(* Logix 5000 project; controller PLC_MCC1300_75F1 vendor 1 type 14 code 166 rev 32.11; software revision 32.04; part 3 of 83 *)
(* tags used below, declared in another part *)
   O : INT[128];
   Z301 : MAC_Zone_ML;

TYPE MAC_TrimmingWheels_PH :
STRUCT
   x0 : BOOL;   // Arming
   x1 : BOOL;
   x2 : BOOL;
   x3 : BOOL;   // Firing operator side
   x4 : BOOL;
   x5 : BOOL;
   x6 : BOOL;   // Firing opposite operator side
   x7 : BOOL;
   x8 : BOOL;
   x9 : BOOL;   // End arming
   x10 : BOOL;
   x11 : BOOL;
   x12 : BOOL;   // End firing
   x13 : BOOL;
   x14 : BOOL;
   x15 : BOOL;   // Stop conveyor request
   x16 : BOOL;
   x17 : BOOL;
   x18 : BOOL;
   x19 : BOOL;
   x20 : BOOL;   // Request position to target
   x21 : BOOL;
   x22 : BOOL;
   x23 : BOOL;   // End position
   x24 : BOOL;
   x25 : BOOL;
   x26 : BOOL;
   x27 : BOOL;
   x28 : BOOL;
   x29 : BOOL;
   x30 : BOOL;
   x31 : BOOL;
END_STRUCT
END_TYPE

TYPE MAC_Zone :
STRUCT
   ST_xConditionOKStopCycle : BOOL;   // Condition OK for stop cycle
   ST_xStartCycleRequest : BOOL;   // Start cycle request
   ST_xCycleON : BOOL;   // Cycle ON
   ST_xStopCycleRequest : BOOL;   // Stop cycle request
   ST_xStopCycleAccepted : BOOL;   // Stop cycle accepted
   ST_xStopCycleReqForAlarms : BOOL;   // Stop cycle request for emergency alarms
   ST_xStopCycleAcptForAlarms : BOOL;   // Stop cycle accepted for emergency alarms
   ST_xConveyorsNotOK : BOOL;   // Conveyors not OK
   ST_xConditionOkPhaseAdvancement : BOOL;   // Condition OK phases advancement
   ST_xConditionOkCycleON : BOOL;   // Condition OK cycle ON
   ST_xConditionOkManualMode : BOOL;   // Condition ok for manual mode
   ST_xCleaningConditionOK : BOOL;   // Cleaning condition OK
   ST_xReqCleaning : BOOL;   // Request cleaning
   ST_xCleaningAccepted : BOOL;   // Cleaning accepted
   ST_xManualModeAccepted : BOOL;   // Manual mode accepted
   ST_xManualModeRequest : BOOL;   // Manual mode request
   ST_xAutoModeAccepted : BOOL;   // Auto mode accepted
   ST_xSelectionManualMode : BOOL;   // Selection manual mode
   ST_xSelectionAutomaticMode : BOOL;   // Selection automatic mode
   ST_xEnableControlError : BOOL;   // Enable control error
   ST_xZoneError : BOOL;   // Zone error
   ST_xAlarmOff : BOOL;   // Alarm OFF
   OSR_xStartCycle : BOOL;   // OSR Start cycle
   OSR_xStopCycle : BOOL;   // OSR Stop cycle
   OSR_xForceStopCycle : BOOL;   // OSR Force stop cycle
   OSR_xAlarmAcoustic : BOOL;   // OSR Alarm acoustic
   OSR_xAlarmMuting : BOOL;   // OSR Alarm muting
   OSR_xAutomaticMode : BOOL;   // OSR Automation mode
   OS_xStartCycle : BOOL;   // OS Start cycle
   OS_xStopCycle : BOOL;   // OS Stop cycle
   OS_xForceStopCycle : BOOL;   // OS Force stop cycle
   OS_xAlarmAcoustic : BOOL;   // OS Alarm acoustic
   OS_xAlarmMuting : BOOL;   // OS Alarm muting
   OS_xAutomaticMode : BOOL;   // OS Automatic mode
   AUX_dSpeedStandby_mm_min : DINT;   // Conveyor speed in stanby [mm/min] (#COSTANT#)
   AUX_dSpeedTINUnload_mm_min : DINT;   // Conveyor speed with stacker in TIM mode [mm/min] (#COSTANT#)
   AUX_dProgressiveID : DINT;   // Progressive ID
   tmON_ResetAlarm : TIMER;   // Reset alarm
   tmON_24Vdc : TIMER;   // Presence 24Vdc timer
   tmON_400Vca : TIMER;   // Presence 400Vca timer
   tmON_EmergencyOK : TIMER;   // Emergency OK timer
   tmON_Cycle : TIMER;   // Cycle ON timer
   tmON_ForceStop : TIMER;   // Force stop cycle timer
   tmON_AllowStopCleaning : TIMER;   // Allow stop cleaning timer
   tmON_CycleAcousticAlarm : TIMER;   // Cycle acoustic alarm timer
END_STRUCT
END_TYPE

TYPE MAC_Zone_ALM :
STRUCT
   rgxEmergency : DINT[3];   // Emergency
   rgxStoppingFault : DINT[1];   // Stopping faults
   rgxFault : DINT[1];   // Faults
   rgxWarning : DINT[2];   // Warning
   rgdFaultCode : DINT[1];   // Fault codes
END_STRUCT
END_TYPE

TYPE MAC_Zone_HMR :
STRUCT
   xZoneAlarm : BOOL;   // Zone alarm
   xCleaningEnabled : BOOL;   // Cleaning enabled
   xSpecialCleaningEnabled : BOOL;   // Special cleaning enabled
   xConsole_M401A_SLTime : BOOL;
   xConsole_M401A_SLAuto : BOOL;
   xConsole_M400A_SL_ManualMode : BOOL;
   dZoneMode : DINT;   // Zone mode (1=Manual 4=Automatic 8=Manual Req)
   dZoneState : DINT;   // Zone status (1=CycleON 2=StopCyc 4=CycleReq 8=StopReq 1024=E-Stop)
   dCabinetState1 : DINT;   // Cabinet status 1 (0=OK; 1=General power alarm; 2=Local power alarm)
   dCabinetState2 : DINT;   // Cabinet status 2 (0=OK; 1=General power alarm; 2=Local power alarm)
   dCleaningState : DINT;   // Cleaning zone status (1=CycleON 2=StopCyc 4=CycleReq 8=StopReq)
   dCleaningSelection : DINT;   // Selection conveyor to start cleaning
   dLineSpeed_mm_min : DINT;   // Line speed [mm/min]
   dSnapSpeed_mm_min : DINT;   // Snap speed [mm/min]
   rgxMan : DINT;   // Manual commands
END_STRUCT
END_TYPE

TYPE MAC_Zone_HMW :
STRUCT
   xManualModeRequest : BOOL;   // Zone manual mode request
   xAutomaticModeRequest : BOOL;   // Zone automatic mode request
   xStartCleanZoneRequest : BOOL;   // Start clean zone request
   xStopCleanZoneRequest : BOOL;   // Stop clean zone request
   xStartCycleRequest : BOOL;   // Start cycle request
   xStopCycleRequest : BOOL;   // Stop cycle request
   xForceStopCycle : BOOL;   // Force stop cycle
   xResetErrorRequest : BOOL;   // Reset error request
   xConsole_SBResetEmergency : BOOL;   // Reset emergency
   xConsole_SB_AlarmOFF : BOOL;   // Acknowledge alarm
   dCleaningSelection : DINT;   // Selection conveyor to start cleaning
   dLocalRemoteSettings : DINT;   // Choose rotate/flip mode from OPT or from Stacker (0=Local "Stacker";1=Remote "OPT")
   dLineSpeed_mm_min : DINT;   // Line speed [mm/min]
   dSnapSpeed_mm_min : DINT;   // Snap speed [mm/min]
   dManualSpeed_mm_min : DINT;   // Manual speed [mm/min]
   rgxMan : DINT;   // Manual commands
END_STRUCT
END_TYPE

TYPE MAC_Zone_ML :
STRUCT
   ST_xSelManuMode : BOOL;   // Selection manual mode
   ST_xSelAutoMode : BOOL;   // Selection auto mode
   ST_xManualModeConditionOK : BOOL;   // Condition Ok for manual mode
   ST_xManuModeReq : BOOL;   // Manual mode request
   ST_xManuModeAccepted : BOOL;   // Manual mode accepted
   ST_xAutoModeAccepted : BOOL;   // Auto mode accepted
   ST_xConditionOKStopCycle : BOOL;   // Condition OK for stop cycle
   ST_xStartCycleRequest : BOOL;   // Start cycle request
   ST_xCycleON : BOOL;   // Cycle ON
   ST_xStopCycleRequest : BOOL;   // Stop cycle request
   ST_xStopCycleAccepted : BOOL;   // Stop cycle accepted
   ST_xStopCycleReqForFaults : BOOL;   // Stop cycle request for stopping faults
   ST_xStopCycleAcceptForFaults : BOOL;   // Stop cycle accepted for stopping faults
   ST_xStopCycleForSaturation : BOOL;   // Stop cycle for saturation on next zone and breaker not available
   ST_xConveyorsNotOK : BOOL;   // Conveyors not OK
   ST_xConditionOkPhaseAdvancement : BOOL;   // Condition OK phases advancement
   ST_xConditionOkCycleON : BOOL;   // Condition OK cycle ON
   ST_xCleaningConditionOK : BOOL;   // Cleaning condition OK
   ST_xZoneReadyForGlass : BOOL;   // Zone ready for glass (enough space to receive glass)
   ST_xReqCleaning : BOOL;   // Request cleaning
   ST_xCleaningAccepted : BOOL;   // Cleaning accepted
   ST_xReqCleaningWrongLength : BOOL;   // Clean cycle request wrong plate length on snap bar
   ST_xReqCleaningMissSnap : BOOL;   // Clean cycle request too many missing snap
   ST_xReqCleaningCPUSwitching : BOOL;   // Clean cycle request for CPU switching
   ST_xReqCleaningBufferOverflow : BOOL;   // Clean cycle for buffer overflow
   ST_xReqCleaningByOperator : BOOL;   // Clean cycle request by operator
   ST_xEnableControlError : BOOL;   // Enable control error
   ST_xZoneError : BOOL;   // Zone error
   ST_xAlarmOff : BOOL;   // Alarm OFF
   ST_xPLC1 : BOOL;   // PLC ID = 1
   ST_xPLC2 : BOOL;   // PLC ID = 2
   ST_xThisPlcActive : BOOL;   // This PLC Active
   ST_xThisPlcActiveForCleaning : BOOL;   // This PLC active for cleaning
   ST_xConditionOkChangeSpeed : BOOL;   // Condition OK for change speed
   ST_rgxConReqClean : DINT;   // Condition request clean
   OSR_xStartCycle : BOOL;   // OSR Start cycle
   OSR_xStopCycle : BOOL;   // OSR Stop cycle
   OSR_xForceStopCycle : BOOL;   // OSR Force stop cycle
   OSR_xAlarmAcoustic : BOOL;   // OSR Alarm acoustic
   OSR_xAlarmMuting : BOOL;   // OSR Alarm muting
   OSR_xThisPlcActive : BOOL;   // OSR ThisPlcActive
   OSR_xLocalCleaningAccepted : BOOL;   // OSR Local cleaning accepted
   OSR_xManualAccepted : BOOL;   // OSR Manual mode accepted
   OSR_xAutoAccepted : BOOL;   // OSR Auto mode accepted
   OS_xStartCycle : BOOL;   // OS Start cycle
   OS_xStopCycle : BOOL;   // OS Stop cycle
   OS_xForceStopCycle : BOOL;   // OS Force stop cycle
   OS_xAlarmAcoustic : BOOL;   // OS Alarm acoustic
   OS_xAlarmMuting : BOOL;   // OS Alarm muting
   OS_xLocalCleaningAccepted : BOOL;   // OS Local cleaning accepted
   OS_xManualAccepted : BOOL;   // OS Manual mode accepted
   OS_xAutoAccepted : BOOL;   // OS Auto mode accepted
   OS_xCleaningAccepted : BOOL;   // OS Cleaning Accepted
   INPUT_x24VdcVoltageON : BOOL;   // 24Vdc Voltage ON
   INPUT_xMainEmergencyON : BOOL;   // Main Emergency ON
   INPUT_xProtectionAirConditioning : BOOL;   // Protection air conditioning
   INPUT_xMCC1201Allow1 : BOOL;   // MCC1201.Allow 1
   INPUT_xMCC1201Allow2 : BOOL;   // MCC1201.Allow 2
   INPUT_xMCC1201Allow3 : BOOL;   // MCC1201.Allow 3
   INPUT_xMCC1201Allow4 : BOOL;   // MCC1201.Allow 4
   INPUT_xCulletAllow1 : BOOL;   // Cullet.Allow 1
   INPUT_xCulletAllow2 : BOOL;   // Cullet.Allow 2
   INPUT_xPowerSupply230V_Service : BOOL;   // Power supply 110/230Vac auxiliary
   INPUT_xPowerSupply230V_PLC1 : BOOL;   // Power supply 110/230Vac PLC1
   INPUT_xPowerSupply230V_PLC2 : BOOL;   // Power supply 110/230Vac PLC2
   INPUT_xPowerSupply24VLogic1 : BOOL;   // Power supply 24Vdc Logic 1
   INPUT_xPowerSupply24VLogic2 : BOOL;   // Power supply 24Vdc Logic 2
   INPUT_xPowerSupply24VLogic3 : BOOL;   // Power supply 24Vdc Logic 3
   INPUT_xPowerSupply24VDrive1 : BOOL;   // Power supply 24Vdc Drive 1
   INPUT_xPowerSupply24VDrive2 : BOOL;   // Power supply 24Vdc Drive 2
   INPUT_xPowerSupply24VDrive3 : BOOL;   // Power supply 24Vdc Drive 3
   INPUT_xPowerSupply400VDrive1 : BOOL;   // Alarm power supply 400/480Vac Drive 1
   INPUT_xPowerSupply400VDrive2 : BOOL;   // Alarm power supply 400/480Vac Drive 2
   INPUT_xPowerSupply400VDrive3 : BOOL;   // Alarm power supply 400/480Vac Drive 3
   INPUT_xPLC_ID_1 : BOOL;   // PLC Identificated as 1
   INPUT_xPLC1Selected : BOOL;   // PLC1 Selected
   INPUT_xPLC2Selected : BOOL;   // PLC2 Selected
   INPUT_xEthernetSwitch24VON : BOOL;   // Ethernet Switch 24Vdc Voltage ON
   INPUT_xEthernetSwitchFault : BOOL;   // Ethernet Switch Fault
   INPUT_xEmergencyLocalization1 : BOOL;   // Emergency localization 1
   INPUT_xEmergencyLocalization2 : BOOL;   // Emergency localization 2
   INPUT_xEmergencyLocalization3 : BOOL;   // Emergency localization 3
   INPUT_xEmergencyLocalization4 : BOOL;   // Emergency localization 4
   INPUT_xEmergencyLocalization5 : BOOL;   // Emergency localization 5
   INPUT_xEmergencyLocalization6 : BOOL;   // Emergency localization 6
   INPUT_xEmergencyLocalization7 : BOOL;   // Emergency localization 7
   INPUT_xEmergencyLocalization8 : BOOL;   // Emergency localization 8
   OUTPUT_xMainEmergencyLamp : BOOL;   // Main emergency ON
   OUTPUT_xMCCSafetyLamp : BOOL;   // Safeties ON
   OUTPUT_xAcousticAlarm : BOOL;   // Acoustic alarm
   OUTPUT_xPLC1Selected : BOOL;   // PLC1 Selected
   OUTPUT_xPLC2Selected : BOOL;   // PLC2 Selected
   OUTPUT_xMCC1201Allow1 : BOOL;   // MCC1201.Allow 1
   OUTPUT_xMCC1201Allow2 : BOOL;   // MCC1201.Allow 2
   OUTPUT_xMCC1201Allow3 : BOOL;   // MCC1201.Allow 3
   OUTPUT_xMCC1201Allow4 : BOOL;   // MCC1201.Allow 4
   OUTPUT_xCulletAllow1 : BOOL;   // Cullet.Allow 1
   OUTPUT_xCulletAllow2 : BOOL;   // Cullet.Allow 2
   OUTPUT_xEmergencyLocalization1 : BOOL;   // Emergency localization 1
   OUTPUT_xEmergencyLocalization2 : BOOL;   // Emergency localization 2
   OUTPUT_xEmergencyLocalization3 : BOOL;   // Emergency localization 3
   OUTPUT_xEmergencyLocalization4 : BOOL;   // Emergency localization 4
   OUTPUT_xEmergencyLocalization5 : BOOL;   // Emergency localization 5
   OUTPUT_xEmergencyLocalization6 : BOOL;   // Emergency localization 6
   AUX_dLehrSpeed_mm_min : DINT;   // Lehr speed [mm/min]
   AUX_dAutoSpeed_mm_min : DINT;   // Automatic speed [mm/min]
   AUX_dSpecialSpeed_mm_min : DINT;   // Special speed [mm/min]
   AUX_dManualSpeed_mm_min : DINT;   // Manual speed [mm/min]
   AUX_dTotalSpaceUsage_cmm : DINT;   // Glass total space usage when goes to next zone [mm/100]
   AUX_dTotalSpaceAvailable_cmm : DINT;   // Conveyor total space available for receive glass in next zone [mm/100]
   AUX_dStartIndexCleaning : DINT;   // Conveyor index of start cleaning
   AUX_dBarPositionCleaning : DINT;   // Progress bar for cleaning position
   tmON_ResetAlarm : TIMER;   // Reset alarm
   tmON_24Vdc : TIMER;   // Presence 24Vdc timer
   tmON_400Vca : TIMER;   // Presence 400Vca timer
   tmON_EmergencyOK : TIMER;   // Emergency OK timer
   tmON_Cycle : TIMER;   // Cycle ON timer
   tmON_ForceStop : TIMER;   // Force stop cycle timer
   tmON_AllowStopCleaning : TIMER;   // Allow stop cleaning timer
   tmON_CycleAcousticAlarm : TIMER;   // Cycle acoustic alarm timer
   tmON_ConveyorsNotOK : TIMER;   // Conveyors not ok
   tmON_StopCycleForFaults : TIMER;   // Stop cycle for stopping faults
   tmON_StopCycleForSaturation : TIMER;   // Enable stop cycle for saturation
END_STRUCT
END_TYPE

TYPE MAC_Zone_ML_ALM :
STRUCT
   rgxEmergency : DINT[3];   // Emergency
   rgxStoppingFault : DINT[1];   // Stopping faults
   rgxFault : DINT[1];   // Faults
   rgxWarning : DINT[1];   // Warning
   rgdFaultCode : DINT[1];   // Fault codes
END_STRUCT
END_TYPE

TYPE MAC_Zone_ML_HMR :
STRUCT
   xZoneAlarm : BOOL;   // Zone fault {x|x|x|x|O}
   xCleaningEnabled : BOOL;   // Cleaning enabled {x|x|x|x|O}
   xChangeThickEnabled : BOOL;   // Thickness change mode enabled {x|x|x|x|O}
   xAutoSpeedAdjustEnabled : BOOL;   // Automatic speed adjustment enabled {x|x|x|x|O}
   rgxConsole_SB : DINT;   // Auxiliary buttons {x|x|x|x|O}
   dZoneMode : DINT;   // Zone mode (1=Manual 4=Automatic 8=Manual Req) {x|x|x|x|O}
   dZoneState : DINT;   // Zone status (1=CycleON 2=StopCyc 4=CycleReq 8=StopReq 1024=E-Stop) {x|x|x|x|O}
   dCabinetState : DINT;   // Cabinet status (0=OK; 1=General power alarm; 2=Local power alarm) {x|x|x|x|O}
   dCleaningState : DINT;   // Cleaning zone status (1=CycleON 2=StopCyc 4=CycleReq 8=StopReq) {x|x|x|x|O}
   dCleaningSelection : DINT;   // Selection conveyor to start cleaning {x|x|x|x|O}
   dAutoSpeedForBreakings_mm_min : DINT;   // dAutoSpeed_mm_min DINT Decimal Automatic speed for breaking zone [mm/min] {mm/min|m/min|x|x|O}
   dAutoSpeed_mm_min : DINT;   // Automatic speed [mm/min] {mm/min|m/min|x|x|O}
   dManualSpeed_mm_min : DINT;   // Manual speed [mm/min] {mm/min|m/min|x|x|O}
   dCleaningEvacuation_cmm : DINT;   // Cleaning evacuation space [mm/100] {mm/100|mm|x|x|O}
   dMinAutoSpeedForBreakings_mm_min : DINT;   // Minimum automatic speed for breaking zone [mm/min] {mm/min|m/min|x|x|O}
   dMinAutoSpeed_mm_min : DINT;   // Minimum automatic speed [mm/min] {mm/min|m/min|x|x|O}
   rSpeedRatioBreakings : REAL;   // Speed ratio for breaking zone (Main line speed/Lehr speed) (Only on 301 zone) {x|x|x|x|O}
   rSpeedRatio : REAL;   // Speed ratio (Main line speed/Lehr speed) {x|x|x|x|O}
   rgxMan : DINT;   // Manual commands {x|x|x|x|O}
   dBarPositionCleaning : DINT;   // Progress bar for cleaning position [mm/100] {mm/100|mm|x|x|O}
END_STRUCT
END_TYPE

TYPE MAC_Zone_ML_HMW :
STRUCT
   xManualModeReq : BOOL;   // Manual mode request {x|x|x|x|O}
   xAutoModeReq : BOOL;   // Automatic mode request {x|x|x|x|O}
   xStartCleanZoneRequest : BOOL;   // Start clean zone request {x|x|x|x|O}
   xStopCleanZoneRequest : BOOL;   // Stop clean zone request {x|x|x|x|O}
   xStartCycleRequest : BOOL;   // Start cycle request {x|x|x|x|O}
   xStopCycleRequest : BOOL;   // Stop cycle request {x|x|x|x|O}
   xForceStopCycle : BOOL;   // Force stop cycle {x|x|x|x|O}
   xResetErrorRequest : BOOL;   // Reset error request {x|x|x|x|O}
   xEnableChangeThick : BOOL;   // Request enable operation in change thickness (Only on 301 zone) {x|x|x|x|O}
   xDisableChangeThick : BOOL;   // Request disable operation in change thickness (Only on 301 zone) {x|x|x|x|O}
   xEnDisableAutoSpeedAdjust : BOOL;   // Automatic speed adjustment enable / disable {x|x|x|x|O}
   rgxConsole_SB : DINT;   // Auxiliary buttons {x|x|x|x|O}
   dCleaningSelection : DINT;   // Selection conveyor to start cleaning (Not for 301 zone) {x|x|x|x|O}
   dSpare : DINT;   // Spare
   dAutoSpeedForBreakings_mm_min : DINT;   // Automatic speed for breaking zone (Only on 301 zone) [mm/min] {mm/min|m/min|7|54|O}
   dAutoSpeed_mm_min : DINT;   // Automatic speed [mm/min] {mm/min|m/min|7|90|O}
   dManualSpeed_mm_min : DINT;   // Manual speed [mm/min] {mm/min|m/min|7|54|O}
   rSpeedRatioBreakings : REAL;   // Speed ratio for breaking zone (Main line speed/Lehr speed) (Only on 301 zone) {x|x|2,0|4,5|O}
   rSpeedRatio : REAL;   // Speed ratio (Main line speed/Lehr speed) {x|x|2,0|4,5|O}
   rgxMan : DINT;   // Manual commands {x|x|x|x|O}
END_STRUCT
END_TYPE

TYPE SpaceConv_Utilities :
STRUCT
   CONST_dSyncMode : DINT;   // Syncrhonization mode [0=No Sync; 1=Sync on head; 2=Sync on tail]
   CONST_dSyncroPhPosition_cmm : DINT;   // Synchronization photocell position [mm/100]
   CONST_dSyncroPhWindow_cmm : DINT;   // Synchronization photocell Windows [mm/100]
   CONST_dConveyorLength_cmm : DINT;   // Conveyor length [mm/100]
   CONST_dConveyorWidth_cmm : DINT;   // Conveyor width [mm/100]
   CONST_dPresetFeedbackTime_ms : DINT;   // Preset feedback Time [ms]
   CONST_rAcceleration_ms2 : REAL;   // Acceleration ramp [m/s2]
   CONST_rDeceleration_ms2 : REAL;   // Deceleration ramp [m/s2]
   CONF_MD1_dScan_ms : DINT;   // Mode1-Previous scan [ms]
   CONF_MD1_xRun : BOOL;   // Mode1-Run
   CONF_MD1_xReverse : BOOL;   // Mode1-Reverse
   CONF_MD1_xTailTracking : BOOL;   // Mode1-Tail tracking active
   CONF_MD1_xHeadTracking : BOOL;   // Mode1-Head tracking active
   CONF_MD2_MD3_dPrstPos_cmm : DINT;   // Mode2|Mode3-Preset position [mm/100]
   CONF_MD4_MD6_dLength_cmm : DINT;   // Mode4|Mode6-Plate length [mm/100]
   CONF_MD7_dOffset_cmm : DINT;   // Mode7-Offset distance between load and unload [mm/100]
   ST_xFeedbackRotation : BOOL;   // Feedback rotation
   ST_xLastModLoadBkw : BOOL;   // Last Modality Load Bkw
   ST_xLastModUnloadBkw : BOOL;   // Last Modality Unload Bkw
   ST_OS_xSynchroPhotocellHead : BOOL;   // OS Sincro Photocel on Head
   ST_OS_xSynchroPhotocellTail : BOOL;   // OS Sincro Photocel on Tail
   ST_dStopLoadForseen_cmm : DINT;   // Stop load forseen [mm/100]
   ST_dRealSpeed_mm_min : DINT;   // Conveyor real speed [mm/min]
   ST_rStepAdvancementH : REAL;   // Step advancement on head [mm/10 per Scan]
   ST_rStepAdvancementT : REAL;   // Step advancement on tail [mm/10 per Scan]
   ST_rSpeedIncrementH_mm_min : REAL;   // Speed increment on head [mm/min]
   ST_rSpeedIncrementT_mm_min : REAL;   // Speed increment on tail [mm/min]
   O_xRampInProgress : BOOL;   // Ramp in progress
   O_xAccInProgress : BOOL;   // Acceleration in progress
   O_xDecInProgress : BOOL;   // Deceleration in progress
   O_xPlateSynchronized : BOOL;   // Plate synchronized
   O_dCountFeedbackTime_ms : DINT;   // Counter feedback time [ms]
   O_dHeadPosition_cmm : DINT;   // Head position [mm/100]
   O_rHeadPosition_cmm : REAL;   // Head position [mm/100]
   O_dTailPosition_cmm : DINT;   // Tail position [mm/100]
   O_rTailPosition_cmm : REAL;   // Tail position [mm/100]
   O_dPresetLoadUnload_cmm : DINT;   // Preset load/unload simultaneously [mm/100]
END_STRUCT
END_TYPE

TYPE UDT_BufferPlate :
STRUCT
   tTracking : UDT_Tracking;
   tData : UDT_ConvoyCap_ZC;
END_STRUCT
END_TYPE

TYPE UDT_Cap :   // Cap data
STRUCT
   dID : DINT;   // Cap ID [Num]
   dProductionID : DINT;   // Cap Production ID [Num]
   dLength_cmm : DINT;   // Cap length [mm/100]
   dWidth_cmm : DINT;   // Cap total width [mm/100]
   dThickness_cmm : DINT;   // Cap thickness [mm/100]
   dGap_cmm : DINT;   // Cap gap between lites [mm/100]
   dIndex : DINT;   // Cap index number in convoy [Num] (0=First cap in convoy)
   dFormat : DINT;   // Plate format [Num] (1=JS 2=LES 3=SSS)
   dNumLites : DINT;   // Number of lites in cap [Num]
   dReqGapForConv_cmm : DINT;   // Request gap between caps for convoy creation [mm/100]
   dMaxCapInConv : DINT;   // Maximum number of caps in convoy [Num]
   dConvTotLength_cmm : DINT;   // Total length of the convoy [mm/100]
   dMinWidth_cmm : DINT;   // Shortest width in use [mm/100]
   dMaxWidth_cmm : DINT;   // Biggest width in use [mm/100]
   dGrossWidth_cmm : DINT;   // Cap gross width [mm/100]
   dNetWidth_cmm : DINT;   // Cap net width [mm/100]
   dDEdgeOpSide_cmm : DINT;   // Double edge dimension - operator side [mm/100]
   dDEdgeOppOpSide_cmm : DINT;   // Double edge dimension - opposite operator side [mm/100]
   dTEdgeOpSide_cmm : DINT;   // Triple edge dimension - operator side [mm/100]
   dTEdgeOppOpSide_cmm : DINT;   // Triple edge dimension - opposite operator side [mm/100]
   dCutWander_cmm : DINT;   // Cap cut wander (- Op. Side + Oppo. Op. Side) [mm/100]
   dNetWander_cmm : DINT;   // Cap net wander (- Op. Side + Oppo. Op. Side) [mm/100]
   dColor : DINT;   // Color code [Num]
   dStackerModality : DINT;   // Stacker Modality [0=MonoPortrait 1=MonoLandscape 10=StereoPortrait 11=StereoLandscape]
   dStackerMode : DINT;   // Stacker Mode [0=Air 1=Tin]
   rgxRequest : DINT;   // Working flag request on cap
   rgxDone : DINT;   // Working flag done on cap
   rgtLite : UDT_Lite[7];
   tFlag : UDT_CapFlags;
END_STRUCT
END_TYPE

TYPE UDT_Cap_SL :   // Cap data
STRUCT
   dID : DINT;   // Cap ID [Num]
   dProductionID : DINT;   // Cap Production ID [Num]
   dLength_cmm : DINT;   // Cap length [mm/100]
   dWidth_cmm : DINT;   // Cap total width [mm/100]
   dThickness_cmm : DINT;   // Cap thickness [mm/100]
   dGap_cmm : DINT;   // Cap gap between lites [mm/100]
   dIndex : DINT;   // Cap index number in convoy [Num] (0=First cap in convoy)
   dFormat : DINT;   // Plate format [Num] (1=JS 2=LES 3=SSS)
   dNumLites : DINT;   // Number of lites in cap [Num]
   dReqGapForConv_cmm : DINT;   // Request gap between caps for convoy creation [mm/100]
   dMaxCapInConv : DINT;   // Maximum number of caps in convoy [Num]
   dConvTotLength_cmm : DINT;   // Total length of the convoy [mm/100]
   dColor : DINT;   // Color code [Num]
   dStackerModality : DINT;   // Stacker Modality [0=MonoPortrait 1=MonoLandscape 10=StereoPortrait 11=StereoLandscape]
   dStackerMode : DINT;   // Stacker Mode [0=Air 1=Tin]
   rgxRequest : DINT;   // Working flag request on cap
   rgxDone : DINT;   // Working flag done on cap
   rgtLite : UDT_Lite_SL[2];
END_STRUCT
END_TYPE

TYPE UDT_CapFlags :   // Cap flags
STRUCT
   xByYCut1 : BOOL;   // Cap done by longitudinal bridge 1
   xByYCut2 : BOOL;   // Cap done by longitudinal bridge 2
   xTrim3OpSide : BOOL;   // Trim 3 Op. Side present (Triple edge)
   xTrim2OpSide : BOOL;   // Trim 2 Op. Side present (Double edge)
   xTrim1OpSide : BOOL;   // Trim 1 Op. Side present (Single edge)
   xTrim1OppOpSide : BOOL;   // Trim 1 Oppo. Op. Side present (Single edge)
   xTrim2OppOpSide : BOOL;   // Trim 2 Oppo. Op. Side present (Double edge)
   xTrim3OppOpSide : BOOL;   // Trim 3 Oppo. Op. Side present (Triple edge)
   rgxIntCut : DINT;   // Internal cuts present between lites ([0]= First cut from Op.Side)
   xOptSelvedgeSel : BOOL;   // Optimizer selvedge selection
   xOptSplitBarSel : BOOL;   // Optimizer split bar selection
   xOptSepRollSel : BOOL;   // Optimizer separator roll selection
   xHookedGeom : BOOL;   // Hooked geometrical camera
   rgxXCutDoneHead : DINT;   // X Cut on head done [Num]
   rgxXCutDoneTail : DINT;   // X Cut on tail [Num]
   rgxYCutHeadDone : DINT;   // Y Cut head done [Mask num]
   tSelvedgeMachine : WorkingFlags_Selvedge;
END_STRUCT
END_TYPE

TYPE UDT_CapsConveyor_ZC :   // Caps tracking conveyor
STRUCT
   xHead : BOOL;   // Head presence on conveyor
   xCenter : BOOL;   // Center presence on conveyor
   xTail : BOOL;   // Tail presence on conveyor
   xPresence : BOOL;   // Plate presence
   dPointer : DINT;   // Head pointer data
   dTailPos_cmm : DINT;   // Tail position [cmm]
   dTailPosConv_cmm : DINT;   // Tail position in conveyor [cmm]
   dCenterPos_cmm : DINT;   // Center position [cmm]
   dCenterPosConv_cmm : DINT;   // Center position in conveyor [cmm]
   dHeadPos_cmm : DINT;   // Head position [cmm]
   dHeadPosConv_cmm : DINT;   // Head position in conveyor [cmm]
   dPresenceHead_cmm : DINT;   // Head position presence [cmm] (the position could be on another conveyor)
   dPresenceTail_cmm : DINT;   // Tail position presence [cmm] (the position could be on another conveyor)
END_STRUCT
END_TYPE

TYPE UDT_Conveyor_Config :
STRUCT
   dLengthConveyor_cmm : DINT;   // Conveyor length [cmm]
   dWidthConveyor_cmm : DINT;   // Conveyor width [cmm]
   dPitchRoller : DINT;   // Conveyor step roller from the next [cmm]
   dMachineIndex : DINT;   // Machine index number for cleaning [Mxxx = xxx*10]
   dZoneConveyor : DINT;   // Conveyor zone belonging [1=xxx1, 2=xxx2, ...]
   dMotorNumber : DINT;   // Motor number [0=single motor, 1=two motors]
   dIndexMainSpeed : DINT;   // Select the conveyor speed [0=AutoSpeed, 1=LehrSpeed, 2=CleaningSpeed, 3=SpecialSpeed, 4=ManualSpeed]
   dGapBetweenM1M2 : DINT;   // Distance between right-left motor
   dSpaceRestartPlate_cmm : DINT;   // Space from previous cap to restart after stop
   dMachineCode : DINT;   // Machine code for Report
   sMachineString : STRING;   // Machine string for Report
   xMotorCmdMainDrive : BOOL;   // Motor command from main drive
   xMotorCmdAndAnomalyInhibit : BOOL;   // Motor command inhibit
   xContinuousConveyor : BOOL;   // Continuous conveyor zone (No saturation with the plate at end of conveyor)
   xWaitNextReadyToMove : BOOL;   // Wait next conveyor ready to move for run
   xWaitGlassForStop : BOOL;   // Continuous conveyor wait glass for for stop zone if there is alarm
   xSimulationMotor : BOOL;   // Simulation motor [0=No simulation, 1=Simulation active]
   xLocalCleaningAllow : BOOL;   // Local cleaning allowed
   xEnableStopPlateContinuousZone : BOOL;   // Enable stop plate in continuous zone
   xOnlyOnePlateAtTheTime : BOOL;   // Access enter new plate - one at the time
   rAccH_ms2 : REAL;   // Acceleration High (for thin glass) [ms2]
   rDecH_ms2 : REAL;   // Deceleration High (for thin glass) [ms2]
   rAccH_s : REAL;   // Acceleration High (for thin glass) [s]
   rDecH_s : REAL;   // Deceleration High (for thin glass) [s]
   rAccL_ms2 : REAL;   // Acceleration Low (for thick glass) [ms2]
   rDecL_ms2 : REAL;   // Deceleration Low (for thick glass) [ms2]
   rAccL_s : REAL;   // Acceleration Low (for thick glass) [s]
   rDecL_s : REAL;   // Deceleration Low (for thick glass) [s]
   rgxAllowedDest : DINT;   // Allowed destinations for scada change after this conveyor
   rgxAllowedCullet : DINT;   // Allowed cullet for scada change after this conveyor
   rgxAllowedQuality : DINT;   // Allowed quality for scada change after this conveyor
END_STRUCT
END_TYPE

TYPE UDT_ConveyorTracking :
STRUCT
   xGlassPresence : BOOL;   // Glass presence on conveyor
   xGlassPresenceOpSide : BOOL;   // Glass presence on conveyor M1
   xGlassPresenceFarSide : BOOL;   // Glass presence on conveyor M2
   xPlatePassagePrevious : BOOL;   // Plate in passage with previous conveyor
   xPlatePassageNext : BOOL;   // Plate in passage with next conveyor
   xGlassPresCom : BOOL;   // Glass presence on conveyor or plate in passage from previous conveyor
   xPlateConvPreviousNext : BOOL;   // Plate in convoy on previous and next conveyor (Internal use)
   xHeadPresenceConv : BOOL;   // Head presence on conveyor
   dStartPosition_cmm : DINT;   // Start position conveyor [cmm]
   dEndPosition_cmm : DINT;   // End position conveyor [cmm]
   dStepAdv_cmm : DINT[2];   // Step advancement [cmm]
   dActualRamp_cmm : DINT[2];   // Actual ramp [cmm]
   dLengthConveyor : DINT;   // Conveyor length [cmm]
   dHeadPosition_cmm : DINT;   // First head position [cmm]
   dTailPosition_cmm : DINT;   // Last tail position [cmm]
   dIndexCaps : DINT;   // Index cap used (Internal use)
   tmON_StopNextConveyor : TIMER;   // Timer for stop next conveyor
   Cap : UDT_CapsConveyor_ZC[10];
END_STRUCT
END_TYPE

TYPE UDT_Convoy_SL :   // Convoy data for load-unload zones
STRUCT
   dLength_cmm : DINT;   // Convoy length [mm/100]
   dTotalCaps : DINT;   // Total caps in convoy [Num] (0=1=No convoy xx=Convoy)
   dGapCaps_cmm : DINT;   // Gap between caps (to next cap) [mm/100]
   dCapIndex : DINT;   // Cap index number in convoy [0 = First cap in convoy]
   dNextCapIndex : DINT;   // Next cap index data (convoy presence) [Num]
   rgtCap : UDT_Cap_SL[2];
   tFlag : UDT_ConvoyFlags;
END_STRUCT
END_TYPE

TYPE UDT_ConvoyCap_ZC :   // Plate data for continuous zones (Tracking circular buffer)
STRUCT
   dLength_cmm : DINT;   // Convoy length [cmm]
   dTotalCaps : DINT;   // Total caps in convoy [Num] (0=1=No convoy xx=Convoy)
   dGapCaps_cmm : DINT;   // Gap between caps (to next cap) [cmm]
   dCapIndex : DINT;   // Cap index number in convoy [0 = First cap in convoy]
   dNextCapIndex : DINT;   // Next cap index data (convoy presence) [Num]
   tFlag : UDT_ConvoyFlags;
   rgtCap : UDT_Cap[1];
   tCapPilkington : DATA_CAP_PILKINGTON;
END_STRUCT
END_TYPE

TYPE UDT_ConvoyFlags :
STRUCT
   tConveyor : WorkingFlags_Conveyor;
   tRotator : WorkingFlags_Rotator;
END_STRUCT
END_TYPE

TYPE UDT_Destination :   // Lite Destinations
STRUCT
   rgxMain : DINT;
   rgxAlternative : DINT;
   rgxSecChoice : DINT;
END_STRUCT
END_TYPE

TYPE UDT_HMI_CAP :   // HMI cap data
STRUCT
   rgtLite : UDT_HMI_LITE[7];   // HMI lite data
END_STRUCT
END_TYPE

TYPE UDT_HMI_LINE_PLATE :
STRUCT
   rgtPlate : UDT_HMI_PLATE[40];   // Scada continuos
END_STRUCT
END_TYPE

TYPE UDT_HMI_LITE :   // HMI Lite data
STRUCT
   dHead_PosX_mm : DINT;   // Plate position X [mm] - Head Position
   dTail_PosX_mm : DINT;   // Plate position X [mm] - Tail Position
   dPlateLength_mm : DINT;   // Plate length [mm]
   dPositionY_mm : DINT;   // Plate position Y [mm]- Operator side
   dPlateWidth_mm : DINT;   // Plate width [mm]
   dPlateId : DINT;   // Plate ID
   dProductionID : DINT;   // Production ID
   dSource : DINT;   // Source
   dDestination : DINT;   // Main destination
   dAlternative : DINT;   // Alternative destination
   dSecondDestination : DINT;   // 2nd choice destination
END_STRUCT
END_TYPE

TYPE UDT_HMI_PLATE :   // HMI Plate data
STRUCT
   rgtCap : UDT_HMI_CAP[1];   // HMI cap data
END_STRUCT
END_TYPE

TYPE UDT_IN_Zone :
STRUCT
   xCleanZoneAccepted : BOOL;   // Zone cleaning accepted
   xExternalConditionCleaning : BOOL;   // External condition for cleaning
   xStartCycleRequest : BOOL;   // Zone start cycle request
   xCycleON : BOOL;   // Cycle ON
   xManualCmdZoneEnabled : BOOL;   // Manual command zone enabled
   xResetFault : BOOL;   // Fault reset
   xCmdFwdAll : BOOL;   // Command forward all
   xCmdBwdAll : BOOL;   // Command backward all
   xEnableControlError : BOOL;   // Enable control error
   dAutoSpeed_mm_min : DINT;   // Automatic speed [mm/min]
   dLehrSpeed_mm_min : DINT;   // Lehr speed [mm/min]
   dCleaningSpeed_mm_min : DINT;   // Cleaning speed [mm/min]
   dSpecialSpeed_mm_min : DINT;   // Special speed [mm/min]
   dManualSpeed_mm_min : DINT;   // Manual speed [mm/min]
   dStartCleaning : DINT;   // Start cleaning conveyor
END_STRUCT
END_TYPE

TYPE UDT_LINE_BUFFER_PLATE :
STRUCT
   rgtPlate : UDT_BufferPlate[40];   // Tracking buffer plate
END_STRUCT
END_TYPE

TYPE UDT_LINE_TRACKING :
STRUCT
   rgtTrkConv : UDT_ConveyorTracking[29];   // Tracking conveyor
END_STRUCT
END_TYPE

TYPE UDT_Lite :   // Lite data
STRUCT
   dID : DINT;   // Lite ID [Num]
   dProductionID : DINT;   // Production ID [Num]
   dQualityID : DINT;   // Quality ID [Num]
   dCameraRecipeID : DINT;   // Camera recipe ID [Num]
   dWidth_cmm : DINT;   // Width [mm/100]
   dBarycenter_cmm : DINT;   // Barycenter [mm/100]
   dCulletCause : DINT;   // Cullet Cause [Num]
   tFlag : UDT_LiteFlags;   // Lite flags
   tDestination : UDT_Destination;   // Destinations of lite
   rgxRequest : DINT;   // Working flag request on lite
   rgxDone : DINT;   // Working flag done on lite
END_STRUCT
END_TYPE

TYPE UDT_Lite_SL :   // Lite data
STRUCT
   dID : DINT;   // Lite ID [Num]
   dProductionID : DINT;   // Production ID [Num]
   dWidth_cmm : DINT;   // Width [mm/100]
   dBarycenter_cmm : DINT;   // Barycenter [mm/100]
   dCulletCause : DINT;   // Cullet Cause [Num]
   tFlag : UDT_LiteFlags;   // Lite flags
   tDestination : UDT_Destination;   // Destinations of lite
   rgxRequest : DINT;   // Working flag request on lite
   rgxDone : DINT;   // Working flag done on lite
END_STRUCT
END_TYPE

TYPE UDT_LiteFlags :   // Lite Flags
STRUCT
   xSaturation : BOOL;   // Saturation lite
   tGeometrical : WorkingFlags_GeomCamera[1];
   tPowder : WorkingFlags_Powder[2];
END_STRUCT
END_TYPE
